      statVarRefList : "LKinLang_typeVarRefList";   // Table containing all variable references
      statLabelList : "LKinLang_typeLabelList";   // Table containing all label references
      statSubPrgList : "LKinLang_typeSubPrgList";   // Table containing all subprogram references
      statStack : "LKinLang_typeStack";   // Static storing for stack elements
      statHierarchicLevel : "LKInLang_typeHierarchicLevel";   // Static storing for hierarchic level info
   END_VAR
   VAR_TEMP
      tempExecute : Bool;   // Temporary value for input 'execute'
      tempStop : Bool;   // Temporary value for input 'stop'
      tempReturnVal : DWord;   // Temporary value for returns of functions
      tempError : Bool;   // Temporary value for error
      tempCounter : Int;   // Temporary counter variable
      tempLabelIndex : Int;   // Temporary counter in labelList
      tempEmptyLineCounter : Int;   // Temporary counter for empty lines / Tenporary counter for empty lines
      tempTokenCounter : Int;   // Temporary counter for token
      tempCycleCounter : Int;   // Temporary value for cycle counter
      tempParseCounter : Int;   // Temporary var to switch direct and follow value parsing
      tempFollowValueCounter : Int;   // Temporary counter for follow values
      tempConditionCounter : Int;   // Temporary counter for conditions
      tempWaitCheckCounter : Int;   // Temporary token counter to check for wait comamnds
      tempFlagOnly : Bool;   // Temporary bit to signalize flag only cmd
      tempWaitTime : Bool;   // Temporary bit to signalize a wait command
      tempAbortRepeat : Bool;   // Temporary bit to abort the repeat loop
      tempParameterIndex : Int;   // Temporary parameter index
      tempSeparatorIndex : Int;   // Temporary separator index
      tempCmdWord : Word;   // Temporary command word
      tempParameterValue : LReal;   // Temporary parameter value
      tempCmdName : String;   // Temporary command name
      tempVarType : Int;   // Temporary variable showing the type of a variable
      tempVarIndex : Int;   // Temporary variable showing the index of a variable
      tempLabelExists : Bool;   // Temporary bit to signalize if a label exists
      tempConditionResult : Bool;   // Temporary result of a condition for conditional jumps
      tempGlobal : Bool;   // Temporary bit to signalize a global variable
      tempPointerOk : Bool;   // Temporary bit to signalize line buffer pointer are ok
      tempLineNumber : UDInt;   // Temporary line number
      tempDelimPos : Array[1..3] of SInt;   // Temporary position of delimiters
      tempTestCommand : "LKinLang_typePathDataElement";   // Temporary PathData command to test iparsed is new
      tempParsedValues : "LKinCtrl_typePathDataElement_advanced";   // Temporary path data element with parsed values
      tempParameterCounter : Array[1.."LKINLANG_MAX_NUMBER_OF_PARAMETERS_PER_LINE"] of "LKinLang_typeParameterCounter";   // Counts the found parameter in one line (G1,F,...)
      tempWaitParameterDefinition : "LKinLang_typeParameterDefinition";   // Temporary definition for a wait command
      tempMathParserResult : "LKinLang_typeMathParserResult";   // Temporary result of the math parser
   END_VAR
   VAR CONSTANT
      MAX_LINES_PER_CYCLE : SInt := 1;   // Maximum lines to be parsed in one call
      MAX_EMPTY_LINES_PER_CYCLE : Int := 5;   // Maximum empty lines handled in one cycle
      MAX_LINES_LABEL_LIST : Int := 5;   // Maximum lines handled in one labelList cycle
      DEFAULT_FLAG_MODE : USInt := 1;   // Flag mode used, if no input default is set
      FB_STATE_NO_PROCESSING : DInt := 0;   // FB state: No processing
      FB_STATE_INIT : DInt := 10;   // FB state: Initialize
      FB_STATE_LOOKUP_PART_1 : DInt := 20;   // FB state: Get commands oart 1
      FB_STATE_LOOKUP_PART_2 : DInt := 21;   // FB state: Get commands part 2
      FB_STATE_PRECHECK_PRG : DInt := 22;   // FB state: Precheck program / FB state: Create label list
      FB_STATE_PARSING : DInt := 30;   // FB state: Parsing
      FB_STATE_STOPPING : DInt := 40;   // FB state: Stopping
      STATE_SEARCH_LINE : Int := 90;   // Internal FB state: Search line in buffer / Internal FB state: Wait until FileHandler has found requested line
      STATE_FILEHANDLER_REQUEST : Int := 91;   // Internal FB state: Wait until FileHandler has found requested line
      STATE_TOKENIZING : Int := 100;   // Internal FB state: Tokenizing
      STATE_INIT_PARSE_LINE : Int := 200;   // Internal FB state: Parsing
      STATE_IS_LINE_VAR_DEF : Int := 201;   // Internal FB state: Is line a variable definition
      STATE_LINE_IS_VAR_DEF : Int := 202;   // Internal FB state: Line is a variable definition
      STATE_IS_LINE_LABEL : Int := 203;   // Internal FB state: Is line a label
      STATE_IS_LINE_GOTO : Int := 204;   // Internal FB state: Is line is jump
      STATE_IS_LINE_STOPRE : Int := 205;   // Internal FB state: Is line a processing stop
      STATE_IS_LINE_IF : Int := 207;   // Internal FB state: Check if line contains IF
      STATE_IS_LINE_WHILE : Int := 208;   // Internal FB state: Check if line contains WHILE
      STATE_IS_LINE_FOR : Int := 209;   // Internal FB state: Check if line contains FOR
      STATE_IS_LINE_SUB : Int := 210;   // Internal FB state: Check if line contains SUB
      STATE_INIT_PARSE_LOOP : Int := 300;   // Internal FB state: Initialize parsing loop
      STATE_IS_TOKEN_SEPARATOR : Int := 310;   // Internal FB state: Check token for separator
      STATE_TOKEN_IS_SEPARATOR : Int := 311;   // Internal FB state: Token is separator
      STATE_IS_TOKEN_NUMBER : Int := 320;   // Internal FB state: Check token for number
      STATE_IS_TOKEN_PARAMETER : Int := 330;   // Internal FB state: Check token for parameter
      STATE_TOKEN_IS_PARAMETER : Int := 331;   // Internal FB state: Token is parameter
      STATE_IS_TOKEN_VARIABLE : Int := 340;   // Internal FB state: Check token for variable
      STATE_TOKEN_IS_VARIABLE : Int := 341;   // Internal FB state: Token is variable
      STATE_TOKEN_IS_UNKNOWN : Int := 350;   // Internal FB state: Token is unknown
      STATE_TOKEN_PROCESSED : Int := 390;   // Internal FB state: Token was processed
      STATE_LINE_PARSED : Int := 400;   // Internal FB state: Parsing single line done
      STATE_CHECK_FOR_NEW_PATH_DATA_CMD : Int := 500;   // Internal FB state: Check parsed command
      STATE_BUILD_PATH_DATA_CMD : Int := 600;   // Internal FB state: Build complete PathData command
      STATE_WRITE_CMD : Int := 700;   // Internal FB state: Write parsed command to path data
      STATE_RESET_AFTER_WRITE : Int := 701;   // Internal FB state: Reset statics and save "old" variables
      STATE_CHECK_END : Int := 800;   // Internal FB state: Check for end of program
      STATE_ERROR : Int := 900;   // Internal FB state: Error
      STATE_PREPROCESSING_STOP : Int := 1000;   // Internal FB state: Wait for MovePath to catch up with execution
      STATUS_EXECUTION_FINISHED : Word := 16#0000;   // Execution finished without errors
      STATUS_NO_CALL : Word := 16#7000;   // No job being currently processed
      STATUS_FIRST_CALL : Word := 16#7001;   // First call after incoming new job (rising edge 'execute')
      STATUS_SUBSEQUENT_CALL : Word := 16#7002;   // Subsequent call during active processing without further details
      STATUS_COMMAND_ABORTED : Word := 16#7FFF;   // Commanded functionality has been aborted by another command
      ERR_UNDEFINED_STATE : Word := 16#8600;   // Error due to an undefined state in state machine
      ERR_PARSING : Word := 16#8601;   // Error while parsing line
      ERR_TOKENIZING : Word := 16#8602;   // Error while tokenizing line
      ERR_LOOKUP : Word := 16#8603;   // Error while creating lookUp table
      ERR_HIERARCHIC_LEVEL_LIST : Word := 16#8604;   // Error while creating hierarchic level list
      ERR_LABEL_LIST : Word := 16#8605;   // Error while creating label list
      ERR_SUB_PROGRAM_LIST : Word := 16#8606;   // Error while creating sub program list
      ERR_LANGUAGE : Word := 16#8200;   // Error missing language definition
      ERR_WRONG_DEFAULTS : Int := -998;   // Error due to missing or wrong default connection
      ERR_LANG_NOT_DEFINED : Int := -999;   // Error selected language not defined
      MINVAL_LREAL : LReal := -1.7976931348623157E+308;   // Minimum value of LREAL
      MAXVAL_LREAL : LReal := 1.7976931348623157E+308;   // Minimum value of LREAL
      MINVAL_DINT : DInt := -2147483648 ;   // Minimum value of DINT
      MAXVAL_DINT : DInt := +2147483647;   // Minimum value of DINT
      MINVAL_INT : Int := -32768;   // Minimum value of INT
      MAXVAL_INT : Int := 32767;   // Maximum vlaue of INT
   END_VAR
BEGIN
   //==========================================================================================
   // SIEMENS AG
   // (c)Copyright 2020 All Rights Reserved
   //------------------------------------------------------------------------------------------
   // Library: LKinLang
   // Tested with: S7-1517T-3 PN/DP
   // Engineering: TIA Portal V15
   // Restrictions: ---
   // Requirements: S7-1500T FW 2.5
   // Functionality: LKinLang_Parser
   // The FB parses strings from line buffer to PathData commands using different language
   // packages.
   // 
   // Support: tech.team.motioncontrol@siemens.com
   // Note: Parameter comments are only available in language 'English (United States)'
   //------------------------------------------------------------------------------------------
   // Change log table:
   // Version    Date          Expert in charge    Changes applied
   // 01.00.00   28.05.2019    FR                  First created version
   // 01.00.01   16.07.2019    FR                  Fixed inserting relative cmd with length 0.0 in some unneccessary cases 
   // 01.00.02   29.07.2019    FR                  Reworked parsing; it is now done directly in this FB
   // 01.01.00   25.11.2019    FR                  Added LRealFlags
   //                                              Added FlagOnlyCmd
   //                                              Added default flag modes as input
   //                                              Fix ignoreAddPointer for LineBuffer
   // 01.01.01   12.02.2020    FR                  Fix circle (auxPoint) recognized as flagOnlyCmd
   // 01.01.02   17.02.2020    FR                  Fix for modal values not taken into account
   //                                              Changed transitionParameter[1] from Int to LReal
   // 01.01.03   17.02.2020    FR                  Changed approach to modal values
   // 01.02.00   15.04.2020    FR                  Added local variables, interface variables and jumps; Added remainingDistance to flagModeDefaults
   // 01.02.01   26.10.2020    FR                  Bugfix when generating label list
   // 01.03.00   01.12.2020    FR                  Added subprograms | Added IF,FOR,WHILE | Several bugfixes
   // 01.03.01   12.04.2021    FR                  Bugfix using followVal for circMode
   //===========================================================================================

   #tempExecute := #execute; // Work with temporary value / create process image
   #tempStop := #stop; // Work with temporary value / create process image

   REGION TRIGGERING
     IF #tempStop = TRUE AND (#statStopOld = FALSE) THEN
       // Stop FB execution
       #statFBState := #FB_STATE_STOPPING;
       // Set status here to avoid return in case of status = NO_CALL
       #statStatus := #STATUS_COMMAND_ABORTED;

     ELSIF (#tempExecute = TRUE) AND (#statExecuteOld = FALSE) AND (#tempStop = FALSE) // Check if FB is triggered
       AND (#statStatus = #STATUS_NO_CALL) // FB must be finished before new job can be started
     THEN // First call; initialize FB
       #statDone := FALSE;
       #statBusy := TRUE;
       #statCommandAborted := FALSE;
       #statError := FALSE;
       #statStatus := #STATUS_FIRST_CALL;

       // Init add pointer (path data)
       #statAddPointer := 0;
       #pathData.pointers.addPointer := 0;
       #pathData.pointers.bufferLocked := TRUE;
       #pathData.pointers.ignoreAddPointer := FALSE;
       #pathData.pointers.preprocessingStop := FALSE;

       // Init retrieve pointer to 0 (line buffer)
       #lineBuffer.pointers.retrievePointer := 0;

       // Reset Error String
       #statErrorString := '';

       // Init look up table
       FOR #tempCounter := 1 TO "LKINLANG_MAX_NUMBER_OF_PARAMETERS" DO
         #statParameterLookUpTable[#tempCounter].parameterNameString := '';
         #statParameterLookUpTable[#tempCounter].parameterNameNumber := 0;
         #statParameterLookUpTable[#tempCounter].parameterNumber := 0;
         #statParameterLookUpTable[#tempCounter].directValueWord := 16#0;
         FOR #tempFollowValueCounter := 1 TO "LKINLANG_NUMBER_OF_FOLLOW_VALUES" DO
           #statParameterLookUpTable[#tempCounter].followValueWords[#tempFollowValueCounter] := 16#0;
         END_FOR;
       END_FOR;

       // FR 2019/04/30
       // Reset path data 
       FOR #tempCounter := 1 TO "LKINCTRL_NO_OF_PATHDATA_ELEMENTS_ADVANCED" DO
         #pathData.commands[#tempCounter] := #statPathDataElementEmpty.pathDataElement;
       END_FOR;

       // Init empty path data element 
       #statModalCommand := #statPathDataElementEmpty;
       #statModalCommandOld := #statPathDataElementEmpty;
       #statModalProgram := #statPathDataElementEmpty;
       #statActualCommand := #statPathDataElementEmpty;
       #statActualCommandOld := #statPathDataElementEmpty;

       #statElementCounter := #statElementCounterEmpty;

       // Init conditions
       FOR #tempCounter := 1 TO "LKINLANG_NUMBER_OF_CONDITIONS" DO
         #statConditionsToCheck[#tempCounter] := #statConditionEmpty;
         #statSetParametersInCmd[#tempCounter] := #statConditionEmpty;
         #statSetParametersInPrg[#tempCounter] := #statConditionEmpty;
       END_FOR;

       // Init tokenized line
       #statTokenizedLine.lineNo := 0;
       #statTokenizedLine.numberOfToken := 0;
       FOR #tempCounter := 1 TO "LKINLANG_MAX_NUMBER_OF_TOKEN_PER_LINE" DO
         #statTokenizedLine.lineToken[#tempCounter] := '';
       END_FOR;

       // Init Positioning mode to absolute
       #statPositioningMode := 1;

       // Init token counter
       #tempTokenCounter := 1;

       // Init condition counter
       #tempConditionCounter := 1;

       // Init flag counter
       #statActualFlagNumber := 0;

       // Init variable definition
       #statVariableDeclaration.localVariables := '';
       #statVariableDeclaration.globalVariables := '';
       #statLocalVariableDefinition.tokenizedString.lineNo := 0;
       #statLocalVariableDefinition.tokenizedString.numberOfToken := 0;
       FOR #tempCounter := 1 TO "LKINLANG_MAX_NUMBER_OF_TOKEN_PER_LINE" DO
         #statLocalVariableDefinition.tokenizedString.lineToken[#tempCounter] := '';
       END_FOR;
       #statLocalVariableDefinition.nameTokenNumber := 0;
       #statLocalVariableDefinition.typeTokenNumber := 0;
       // Init global
       #statGlobalVariableDefinition := #statLocalVariableDefinition;


       // Init vars & counter
       FOR #tempVarIndex := 1 TO "LKINLANG_NUMBER_OF_LOCAL_BOOL" DO
         #statVariables.boolean[#tempVarIndex] := FALSE;
       END_FOR;
       FOR #tempVarIndex := 1 TO "LKINLANG_NUMBER_OF_LOCAL_DINT" DO
         #statVariables.dints[#tempVarIndex] := 0;
       END_FOR;
       FOR #tempVarIndex := 1 TO "LKINLANG_NUMBER_OF_LOCAL_LREAL" DO
         #statVariables.lreals[#tempVarIndex] := 0.0;
       END_FOR;
       #statVariables.boolCounter := 0;
       #statVariables.dintCounter := 0;
       #statVariables.lrealCounter := 0;

       // Remove local vars from var ref table
       FOR #tempVarIndex := 1 TO "LKINLANG_NUMBER_OF_VAR_REFS" DO
         IF #statVarRefList.references[#tempVarIndex].type < "LKINLANG_VAR_TYPE_INTERFACE_BOOL" THEN
           #statVarRefList.references[#tempVarIndex].index := 0;
           #statVarRefList.references[#tempVarIndex].name := '';
           #statVarRefList.references[#tempVarIndex].type := 0;
           #statVarRefList.references[#tempVarIndex].scope := 0;
         END_IF;
       END_FOR;

       // Reset number of references
       #statVarRefList.numberOfReferences := 0;

       // Reset LabelList
       FOR #tempCounter := 1 TO "LKINLANG_NUMBER_OF_LABELS" DO
         #statLabelList.labels[#tempCounter].labelName := '';
         #statLabelList.labels[#tempCounter].lineNumber := 0;
         #statLabelList.labels[#tempCounter].hierarchicLevel := 0;
       END_FOR;
       #statLabelList.numberOfLabels := 0;

       // Reset hierarchicLevel
       FOR #tempCounter := 1 TO "LKINLANG_NUMBER_OF_HIERARCHICLEVEL" DO
         #statHierarchicLevel.levels[#tempCounter].level := 0;
         #statHierarchicLevel.levels[#tempCounter].lineNumber := 0;
         #statHierarchicLevel.levels[#tempCounter].type := 0;
       END_FOR;
       #statHierarchicLevel.numberOfLevels := 0;
       #statHierarchicLevel.currentLevel := 0;

       // Reset Stack
       FOR #tempCounter := 1 TO "LKINLANG_NUMBER_OF_STACK_ELEMENTS" DO
         #statStack.stackElements[#tempCounter].lineNumberStart := 0;
         #statStack.stackElements[#tempCounter].lineNumberEnd := 0;
         #statStack.stackElements[#tempCounter].type := 0;
         #statStack.stackElements[#tempCounter].increment := 0;
         #statStack.stackElements[#tempCounter].quantity := 0;
         #statStack.stackElements[#tempCounter].variableRef.index := 0;
         #statStack.stackElements[#tempCounter].variableRef.type := 0;
         #statStack.stackElements[#tempCounter].variableRef.name := '';
       END_FOR;
       #statStack.numberOfElements := 0;

       // Reset subprogram list
       FOR #tempCounter := 1 TO "LKINLANG_NUMBER_OF_SUBPROGRAMS" DO
         #statSubPrgList.subPrgs[#tempCounter].prgName := '';
         #statSubPrgList.subPrgs[#tempCounter].lineNumberStart := 0;
         #statSubPrgList.subPrgs[#tempCounter].lineNumberEnd := 0;
       END_FOR;
       #statSubPrgList.numberOfSubPrgs := 0;

       // Reset parameter definition
       #statParameterDefinition := #statParameterDefinitionEmpty;

       // Select Language
       #statSelectedLanguage := #language;

       // Syntax check
       #statSyntaxCheck := #syntaxCheck;

       // Reset stringExpression
       #statStringExpression := '';

       // Reset requested line
       #statSearchedLine := 0;

       // Set file state initially
       IF #lineBuffer.info.fileState = "LKINLANG_FILE_STATE_LOADING" THEN
         #lineBuffer.info.fileState := "LKINLANG_FILE_STATE_RUNNING_LOADING";
       ELSE
         #lineBuffer.info.fileState := "LKINLANG_FILE_STATE_RUNNING";
       END_IF;

       // State machine - start processing
       #statFBState := #FB_STATE_INIT;

     ELSIF (#statStatus = #STATUS_FIRST_CALL) THEN
       #statStatus := #STATUS_SUBSEQUENT_CALL;
     END_IF;

     // Edge detection 'execute' input
     #statExecuteOld := #tempExecute;
     // Edge detection 'stop' input
     #statStopOld := #tempStop;
   END_REGION TRIGGERING

   IF (#statStatus = #STATUS_NO_CALL) THEN // Nothing to do -> End here to reduce "system load"
     RETURN;
   END_IF;

   REGION STATE_MACHINE
     CASE #statFBState OF // State machine of FB
       #FB_STATE_NO_PROCESSING: // No processing active (Note: this state must always be present and left empty)
         ;

         // ------------------------------------------------------------------------------------------
         // Get separators, mergers and valid counts from language and save in static arrays
         // ------------------------------------------------------------------------------------------  
       #FB_STATE_INIT:
         REGION FB_STATE_INIT
           // Get separators and mergers from language package
           #tempParameterIndex := -1;
           "LKinLang_SelectLangPackage"(language := #statSelectedLanguage,
                                        variableDeclarations => #statVariableDeclaration,
                                        keyToken => #statKeyToken,
                                        parameterDefinition := #statParameterDefinition,
                                        separators => #statSeparators,
                                        mergers => #statMergers,
                                        validCounts => #statValidCounts,
                                        parameterNumber := #tempParameterIndex,
                                        parameterDefaults := #parameterDefaults);

           IF #tempParameterIndex = #ERR_LANG_NOT_DEFINED THEN
             // Error language not defined
             #statStatus := #ERR_LANGUAGE;
             #statStateIntern := #STATE_ERROR;
             #statErrorString := CONCAT(IN1 := #statErrorString, IN2 := 'Error: Selected language ');
             #statErrorString := CONCAT(IN1 := #statErrorString, IN2 := INT_TO_STRING(#statSelectedLanguage));
             #statErrorString := CONCAT(IN1 := #statErrorString, IN2 := ' not defined');
           END_IF;

           IF #tempParameterIndex = #ERR_WRONG_DEFAULTS THEN
             // Error language not defined
             #statStatus := #ERR_LANGUAGE;
             #statStateIntern := #STATE_ERROR;
             #statErrorString := CONCAT(IN1 := #statErrorString, IN2 := 'Error: Type of parameter defaults not matching language');
           END_IF;

           #statLastIndexOfMerger := 1;

           // Search last entry in mergers to save time in tokenizing
           FOR #tempCounter := 1 TO "LKINLANG_NUMBER_OF_MERGERS" DO
             IF #statMergers[#tempCounter] <> 16#00 THEN
               #statLastIndexOfMerger := #tempCounter;
             END_IF;
           END_FOR;

           // Tokenize variable definition string from language package
           #tempReturnVal := "LKinLang_TokenizeSlot"(lastIndexOfMerger := #statLastIndexOfMerger,
                                                     lineNumber := 0,
                                                     line := #statVariableDeclaration.localVariables,
                                                     separators := #statSeparators,
                                                     mergers := #statMergers,
                                                     preprocessorConfig := #preProcessConfig,
                                                     tokenizedLine => #statLocalVariableDefinition.tokenizedString,
                                                     errorString := #statErrorString);

           // Search tokenized variable definiton for name and type token
           FOR #tempCounter := 1 TO #statLocalVariableDefinition.tokenizedString.numberOfToken DO
             IF #statLocalVariableDefinition.tokenizedString.lineToken[#tempCounter] = '_name_' THEN
               #statLocalVariableDefinition.nameTokenNumber := DINT_TO_USINT(#tempCounter);
             ELSIF #statLocalVariableDefinition.tokenizedString.lineToken[#tempCounter] = '_type_' THEN
               #statLocalVariableDefinition.typeTokenNumber := DINT_TO_USINT(#tempCounter);
             END_IF;
           END_FOR;

           // Double check 
           IF #statLocalVariableDefinition.nameTokenNumber = 0
             OR #statLocalVariableDefinition.typeTokenNumber = 0 THEN
             // Error no valid variable definition found
             #statStatus := #ERR_LANGUAGE;
             #statStateIntern := #STATE_ERROR;
             #statErrorString := CONCAT(IN1 := #statErrorString, IN2 := 'Error: No valid variable definition found');
           END_IF;

           // Tokenize variable definition string from language package
           #tempReturnVal := "LKinLang_TokenizeSlot"(lastIndexOfMerger := #statLastIndexOfMerger,
                                                     lineNumber := 0,
                                                     line := #statVariableDeclaration.globalVariables,
                                                     separators := #statSeparators,
                                                     mergers := #statMergers,
                                                     preprocessorConfig := #preProcessConfig,
                                                     tokenizedLine => #statGlobalVariableDefinition.tokenizedString,
                                                     errorString := #statErrorString);

           // Search tokenized variable definiton for name and type token
           FOR #tempCounter := 1 TO #statGlobalVariableDefinition.tokenizedString.numberOfToken DO
             IF #statGlobalVariableDefinition.tokenizedString.lineToken[#tempCounter] = '_name_' THEN
               #statGlobalVariableDefinition.nameTokenNumber := DINT_TO_USINT(#tempCounter);
             ELSIF #statGlobalVariableDefinition.tokenizedString.lineToken[#tempCounter] = '_type_' THEN
               #statGlobalVariableDefinition.typeTokenNumber := DINT_TO_USINT(#tempCounter);
             END_IF;
           END_FOR;

           // Double check 
           IF #statGlobalVariableDefinition.nameTokenNumber = 0
             OR #statGlobalVariableDefinition.typeTokenNumber = 0 THEN
             // Error no valid variable definition found
             #statStatus := #ERR_LANGUAGE;
             #statStateIntern := #STATE_ERROR;
             #statErrorString := CONCAT(IN1 := #statErrorString, IN2 := 'Error: No valid variable definition found');
           END_IF;

           // Check syntax check mode
           IF #statSyntaxCheck <> "LKINLANG_SYNTAX_CHECK_AND_EXECUTE"
             AND #statSyntaxCheck <> "LKINLANG_SYNTAX_CHECK_OFF"
             AND #statSyntaxCheck <> "LKINLANG_SYNTAX_CHECK_ONLY" THEN
             // Error no valid syntax check mode
             #statStatus := #ERR_LANGUAGE;
             #statStateIntern := #STATE_ERROR;
             #statErrorString := CONCAT(IN1 := #statErrorString, IN2 := 'Error: No valid syntax check setting');
           END_IF;

           // Next state
           #statFBState := #FB_STATE_LOOKUP_PART_1;
         END_REGION FB_STATE_INIT

         // ------------------------------------------------------------------------------------------
         // Get first part of language definition where ParameterNameNumber <> -1 
         // Save the parameter numbers in lookup-table
         // The lookup-table is later used while parsing to have faster access to the parameter definition
         // ------------------------------------------------------------------------------------------ 
       #FB_STATE_LOOKUP_PART_1:
         REGION FB_STATE_LOOKUP_PART_1
           // Init command counter
           #statLookUpTableCounter := 1;

           // Get commands with parameterNameNumber <> -1
           "LKinLang_CreateParameterLookUpTable"(language := #statSelectedLanguage,
                                                 mode := 0, //  ParameterNameNumber <> -1
                                                 error => #tempError,
                                                 lastIndexLookUp => #statLastIndexLookUp,
                                                 parameterLookUpTable := #statParameterLookUpTable,
                                                 parameterDefaults := #parameterDefaults,
                                                 parameterCounter := #statLookUpTableCounter,
                                                 errorString := #statErrorString);
           IF #tempError THEN
             // Error while creating look up table --> Exit
             #statStatus := #ERR_LOOKUP;
             #statStateIntern := #STATE_ERROR;
           ELSE
             // Next state
             #statFBState := #FB_STATE_LOOKUP_PART_2;
           END_IF;
         END_REGION FB_STATE_LOOKUP_PART_1

         // ------------------------------------------------------------------------------------------
         // Get second part of language definition where ParameterNameNumber = -1 
         // Save the parameter numbers in lookup-table
         // Initialize internal states (IF cases)
         // ------------------------------------------------------------------------------------------ 
       #FB_STATE_LOOKUP_PART_2:
         REGION FB_STATE_LOOKUP_PART_2
           // Get commands with parameterNameNumber = -1
           "LKinLang_CreateParameterLookUpTable"(language := #statSelectedLanguage,
                                                 mode := 1, // ParameterNameNumber = -1
                                                 error => #tempError,
                                                 lastIndexLookUp => #statLastIndexLookUp,
                                                 parameterLookUpTable := #statParameterLookUpTable,
                                                 parameterDefaults := #parameterDefaults,
                                                 parameterCounter := #statLookUpTableCounter,
                                                 errorString := #statErrorString);
           IF #tempError THEN
             // Error while creating look up table --> Exit
             #statStatus := #ERR_LOOKUP;
             #statStateIntern := #STATE_ERROR;
           ELSE
             // Next state
             //#statFBState := #FB_STATE_PARSING;
             #statFBState := #FB_STATE_PRECHECK_PRG;

             // Set internal state to tokenizing
             #statStateIntern := #STATE_TOKENIZING;
           END_IF;
         END_REGION FB_STATE_LOOKUP_PART_2

         // ------------------------------------------------------------------------------------------
         // Here the whole program is checked
         // Following things should be done here:
         // - Get HierarchicLevel
         // - Create Label List
         // - Get ProgramName (PRG)?
         // - Get SubProgram List
         // - Check for M17/M30?
         //  
         // After all this is done without error, the actual parsing can be started 
         // The filehandler must be restarted and the lineBuffer must be reset
         // then switch over to FB state "PARSING"
         // The tokenization has to be done here and in state PARSING --> Maybe find a better solution?
         // ------------------------------------------------------------------------------------------
       #FB_STATE_PRECHECK_PRG:
         REGION FB_STATE_PRECHECK_PRG
           // Reset empty line counter
           #tempEmptyLineCounter := 0;

           // Repeat tokenizing until aborted
           // Aborted by:
           // - No new lines in line buffer
           // - End of file reached
           REPEAT

             // Check lineBuffer pointer if next line can be retrieved
             IF ((#lineBuffer.pointers.addPointer > #lineBuffer.pointers.retrievePointer
               AND NOT #lineBuffer.pointers.bufferLocked // Buffer is not locked by fileHandler
               AND NOT #lineBuffer.pointers.addPointerRestarted) // Overflow of ring buffer
               OR
               (#lineBuffer.pointers.addPointer < #lineBuffer.pointers.retrievePointer
               AND #lineBuffer.pointers.addPointerRestarted
               AND NOT #lineBuffer.pointers.bufferLocked))
               OR #lineBuffer.pointers.ignoreAddPointer // FR 25.11.2019
             THEN

               // Increment retrieve pointer
               IF #lineBuffer.pointers.retrievePointer < "LKINLANG_LAST_INDEX_LINE_BUFFER" THEN
                 #lineBuffer.pointers.retrievePointer += 1;

                 // Reset retrieve pointer to 1 and reset overflow variable
               ELSIF #lineBuffer.pointers.retrievePointer >= "LKINLANG_LAST_INDEX_LINE_BUFFER" THEN
                 #lineBuffer.pointers.retrievePointer := 1;
                 #lineBuffer.pointers.addPointerRestarted := FALSE;
               END_IF;

               // ------------------------------------------------------------------------------------------
               // Get hierarchic level
               // ------------------------------------------------------------------------------------------
               // Get hierarchic level --> Check for IF;WHILE;FOR and increse or decrease level
               // Hierarchic level is needed to check if jumps are allowed
               REGION GET_HIERARCHIC_LEVEL
                 // Check if line contains IF token
                 IF FIND(IN1 := #lineBuffer.lines[#lineBuffer.pointers.retrievePointer].content, IN2 := #statKeyToken.tokenIf) <> 0 THEN
                   // Tokenize line where retrieve pointer is pointing at
                   #tempReturnVal := "LKinLang_TokenizeSlot"(lastIndexOfMerger := #statLastIndexOfMerger,
                                                             lineNumber := #lineBuffer.lines[#lineBuffer.pointers.retrievePointer].number,
                                                             line := #lineBuffer.lines[#lineBuffer.pointers.retrievePointer].content,
                                                             separators := #statSeparators,
                                                             mergers := #statMergers,
                                                             preprocessorConfig := #preProcessConfig,
                                                             tokenizedLine => #statTokenizedLine,
                                                             errorString := #statErrorString);

                   // Check if line has content
                   IF #statTokenizedLine.numberOfToken > 0 THEN
                     // Check if line starts with IF token
                     IF #statTokenizedLine.lineToken[#statTokenizedLine.numberOfToken] = #statKeyToken.tokenIf THEN
                       // Increase array index
                       #statHierarchicLevel.numberOfLevels += 1;
                       // Check if index is ok
                       IF #statHierarchicLevel.numberOfLevels <= "LKINLANG_NUMBER_OF_HIERARCHICLEVEL" THEN
                         // Increase hierarchic level
                         #statHierarchicLevel.currentLevel += 1;
                         // Store entry
                         #statHierarchicLevel.levels[#statHierarchicLevel.numberOfLevels].level := #statHierarchicLevel.currentLevel;
                         #statHierarchicLevel.levels[#statHierarchicLevel.numberOfLevels].lineNumber := #statTokenizedLine.lineNo;
                         #statHierarchicLevel.levels[#statHierarchicLevel.numberOfLevels].type := "LKINLANG_ENTRY_TYPE_IF"; // Type for IF
                       ELSE
                         // Error hierarchic level array overflow
                         #statStatus := #ERR_HIERARCHIC_LEVEL_LIST;
                         #statStateIntern := #STATE_ERROR;
                         #statErrorString := CONCAT(IN1 := #statErrorString, IN2 := 'Error: Maximum array index of hierarchic level reached');
                         #statErrorString := CONCAT(IN1 := #statErrorString, IN2 := ' in line: ');
                         #statErrorString := CONCAT(IN1 := #statErrorString, IN2 := UDINT_TO_STRING(#statTokenizedLine.lineNo));
                       END_IF;
                     END_IF;
                   END_IF;
                 END_IF;

                 // Check if line contains ELSE token
                 IF FIND(IN1 := #lineBuffer.lines[#lineBuffer.pointers.retrievePointer].content, IN2 := #statKeyToken.tokenElse) <> 0 THEN
                   // Tokenize line where retrieve pointer is pointing at
                   #tempReturnVal := "LKinLang_TokenizeSlot"(lastIndexOfMerger := #statLastIndexOfMerger,
                                                             lineNumber := #lineBuffer.lines[#lineBuffer.pointers.retrievePointer].number,
                                                             line := #lineBuffer.lines[#lineBuffer.pointers.retrievePointer].content,
                                                             separators := #statSeparators,
                                                             mergers := #statMergers,
                                                             preprocessorConfig := #preProcessConfig,
                                                             tokenizedLine => #statTokenizedLine,
                                                             errorString := #statErrorString);

                   // Check if line has content
                   IF #statTokenizedLine.numberOfToken > 0 THEN
                     // Check if line starts with ELSE token
                     IF #statTokenizedLine.lineToken[#statTokenizedLine.numberOfToken] = #statKeyToken.tokenElse THEN
                       // Check if number of token is exactly 1 --> Nothing more allowed
                       IF #statTokenizedLine.numberOfToken = 1 THEN
                         // Increase array index
                         #statHierarchicLevel.numberOfLevels += 1;
                         // Check if index is ok
                         IF #statHierarchicLevel.numberOfLevels <= "LKINLANG_NUMBER_OF_HIERARCHICLEVEL" THEN
                           // Level does not change
                           // Store entry
                           #statHierarchicLevel.levels[#statHierarchicLevel.numberOfLevels].level := #statHierarchicLevel.currentLevel;
                           #statHierarchicLevel.levels[#statHierarchicLevel.numberOfLevels].lineNumber := #statTokenizedLine.lineNo;
                           #statHierarchicLevel.levels[#statHierarchicLevel.numberOfLevels].type := "LKINLANG_ENTRY_TYPE_ELSE"; // Type for ELSE
                         ELSE
                           // Error hierarchic level array overflow
                           #statStatus := #ERR_HIERARCHIC_LEVEL_LIST;
                           #statStateIntern := #STATE_ERROR;
                           #statErrorString := CONCAT(IN1 := #statErrorString, IN2 := 'Error: Maximum array index of hierarchic level reached');
                           #statErrorString := CONCAT(IN1 := #statErrorString, IN2 := ' in line: ');
                           #statErrorString := CONCAT(IN1 := #statErrorString, IN2 := UDINT_TO_STRING(#statTokenizedLine.lineNo));
                         END_IF;
                       ELSE
                         // Error wrong usage of ELSE
                         #statStatus := #ERR_HIERARCHIC_LEVEL_LIST;
                         #statStateIntern := #STATE_ERROR;
                         #statErrorString := CONCAT(IN1 := #statErrorString, IN2 := 'Error: Wrong syntax of ');
                         #statErrorString := CONCAT(IN1 := #statErrorString, IN2 := #statKeyToken.tokenElse);
                         #statErrorString := CONCAT(IN1 := #statErrorString, IN2 := ' in line: ');
                         #statErrorString := CONCAT(IN1 := #statErrorString, IN2 := UDINT_TO_STRING(#statTokenizedLine.lineNo));
                       END_IF;
                     END_IF;
                   END_IF;
                 END_IF;

                 // Check if line contains ENDIF token
                 IF FIND(IN1 := #lineBuffer.lines[#lineBuffer.pointers.retrievePointer].content, IN2 := #statKeyToken.tokenEndIf) <> 0 THEN
                   // Tokenize line where retrieve pointer is pointing at
                   #tempReturnVal := "LKinLang_TokenizeSlot"(lastIndexOfMerger := #statLastIndexOfMerger,
                                                             lineNumber := #lineBuffer.lines[#lineBuffer.pointers.retrievePointer].number,
                                                             line := #lineBuffer.lines[#lineBuffer.pointers.retrievePointer].content,
                                                             separators := #statSeparators,
                                                             mergers := #statMergers,
                                                             preprocessorConfig := #preProcessConfig,
                                                             tokenizedLine => #statTokenizedLine,
                                                             errorString := #statErrorString);

                   // Check if line has content
                   IF #statTokenizedLine.numberOfToken > 0 THEN
                     // Check if line starts with ENDIF token
                     IF #statTokenizedLine.lineToken[#statTokenizedLine.numberOfToken] = #statKeyToken.tokenEndIf THEN
                       // Check if number of token is exactly 1 --> Nothing more allowed
                       IF #statTokenizedLine.numberOfToken = 1 THEN
                         // Increase array index
                         #statHierarchicLevel.numberOfLevels += 1;
                         // Check if index is ok
                         IF #statHierarchicLevel.numberOfLevels <= "LKINLANG_NUMBER_OF_HIERARCHICLEVEL" THEN
                           // Store entry
                           #statHierarchicLevel.levels[#statHierarchicLevel.numberOfLevels].level := #statHierarchicLevel.currentLevel;
                           #statHierarchicLevel.levels[#statHierarchicLevel.numberOfLevels].lineNumber := #statTokenizedLine.lineNo;
                           #statHierarchicLevel.levels[#statHierarchicLevel.numberOfLevels].type := "LKINLANG_ENTRY_TYPE_ENDIF"; // Type for ENDIF

                           // Decrease hierarchic level
                           #statHierarchicLevel.currentLevel -= 1;
                         ELSE
                           // Error hierarchic level array overflow
                           #statStatus := #ERR_HIERARCHIC_LEVEL_LIST;
                           #statStateIntern := #STATE_ERROR;
                           #statErrorString := CONCAT(IN1 := #statErrorString, IN2 := 'Error: Maximum array index of hierarchic level reached');
                           #statErrorString := CONCAT(IN1 := #statErrorString, IN2 := ' in line: ');
                           #statErrorString := CONCAT(IN1 := #statErrorString, IN2 := UDINT_TO_STRING(#statTokenizedLine.lineNo));
                         END_IF;
                       ELSE
                         // Error wrong usage of ENDIF
                         #statStatus := #ERR_HIERARCHIC_LEVEL_LIST;
                         #statStateIntern := #STATE_ERROR;
                         #statErrorString := CONCAT(IN1 := #statErrorString, IN2 := 'Error: Wrong syntax of ');
                         #statErrorString := CONCAT(IN1 := #statErrorString, IN2 := #statKeyToken.tokenEndIf);
                         #statErrorString := CONCAT(IN1 := #statErrorString, IN2 := ' in line: ');
                         #statErrorString := CONCAT(IN1 := #statErrorString, IN2 := UDINT_TO_STRING(#statTokenizedLine.lineNo));
                       END_IF;
                     END_IF;
                   END_IF;
                 END_IF;

                 // Check if line contains WHILE token
                 IF FIND(IN1 := #lineBuffer.lines[#lineBuffer.pointers.retrievePointer].content, IN2 := #statKeyToken.tokenWhile) <> 0 THEN
                   // Tokenize line where retrieve pointer is pointing at
                   #tempReturnVal := "LKinLang_TokenizeSlot"(lastIndexOfMerger := #statLastIndexOfMerger,
                                                             lineNumber := #lineBuffer.lines[#lineBuffer.pointers.retrievePointer].number,
                                                             line := #lineBuffer.lines[#lineBuffer.pointers.retrievePointer].content,
                                                             separators := #statSeparators,
                                                             mergers := #statMergers,
                                                             preprocessorConfig := #preProcessConfig,
                                                             tokenizedLine => #statTokenizedLine,
                                                             errorString := #statErrorString);

                   // Check if line has content
                   IF #statTokenizedLine.numberOfToken > 0 THEN
                     // Check if line starts with WHILE token
                     IF #statTokenizedLine.lineToken[#statTokenizedLine.numberOfToken] = #statKeyToken.tokenWhile THEN
                       // Increase array index
                       #statHierarchicLevel.numberOfLevels += 1;
                       // Check if index is ok
                       IF #statHierarchicLevel.numberOfLevels <= "LKINLANG_NUMBER_OF_HIERARCHICLEVEL" THEN
                         // Increase hierarchic level
                         #statHierarchicLevel.currentLevel += 1;
                         // Store entry
                         #statHierarchicLevel.levels[#statHierarchicLevel.numberOfLevels].level := #statHierarchicLevel.currentLevel;
                         #statHierarchicLevel.levels[#statHierarchicLevel.numberOfLevels].lineNumber := #statTokenizedLine.lineNo;
                         #statHierarchicLevel.levels[#statHierarchicLevel.numberOfLevels].type := "LKINLANG_ENTRY_TYPE_WHILE"; // Type for WHILE
                       ELSE
                         // Error hierarchic level array overflow
                         #statStatus := #ERR_HIERARCHIC_LEVEL_LIST;
                         #statStateIntern := #STATE_ERROR;
                         #statErrorString := CONCAT(IN1 := #statErrorString, IN2 := 'Error: Maximum array index of hierarchic level reached');
                         #statErrorString := CONCAT(IN1 := #statErrorString, IN2 := ' in line: ');
                         #statErrorString := CONCAT(IN1 := #statErrorString, IN2 := UDINT_TO_STRING(#statTokenizedLine.lineNo));
                       END_IF;
                     END_IF;
                   END_IF;
                 END_IF;

                 // Check if line contains ENDWHILE token
                 IF FIND(IN1 := #lineBuffer.lines[#lineBuffer.pointers.retrievePointer].content, IN2 := #statKeyToken.tokenEndWhile) <> 0 THEN
                   // Tokenize line where retrieve pointer is pointing at
                   #tempReturnVal := "LKinLang_TokenizeSlot"(lastIndexOfMerger := #statLastIndexOfMerger,
                                                             lineNumber := #lineBuffer.lines[#lineBuffer.pointers.retrievePointer].number,
                                                             line := #lineBuffer.lines[#lineBuffer.pointers.retrievePointer].content,
                                                             separators := #statSeparators,
                                                             mergers := #statMergers,
                                                             preprocessorConfig := #preProcessConfig,
                                                             tokenizedLine => #statTokenizedLine,
                                                             errorString := #statErrorString);

                   // Check if line has content
                   IF #statTokenizedLine.numberOfToken > 0 THEN
                     // Check if line starts with ENDWHILE token
                     IF #statTokenizedLine.lineToken[#statTokenizedLine.numberOfToken] = #statKeyToken.tokenEndWhile THEN
                       // Check if number of token is exactly 1 --> Nothing more allowed
                       IF #statTokenizedLine.numberOfToken = 1 THEN
                         // Increase array index
                         #statHierarchicLevel.numberOfLevels += 1;
                         // Check if index is ok
                         IF #statHierarchicLevel.numberOfLevels <= "LKINLANG_NUMBER_OF_HIERARCHICLEVEL" THEN
                           // Store entry
                           #statHierarchicLevel.levels[#statHierarchicLevel.numberOfLevels].level := #statHierarchicLevel.currentLevel;
                           #statHierarchicLevel.levels[#statHierarchicLevel.numberOfLevels].lineNumber := #statTokenizedLine.lineNo;
                           #statHierarchicLevel.levels[#statHierarchicLevel.numberOfLevels].type := "LKINLANG_ENTRY_TYPE_ENDWHILE"; // Type for ENDWHILE

                           // Decrease hierarchic level
                           #statHierarchicLevel.currentLevel -= 1;
                         ELSE
                           // Error hierarchic level array overflow
                           #statStatus := #ERR_HIERARCHIC_LEVEL_LIST;
                           #statStateIntern := #STATE_ERROR;
                           #statErrorString := CONCAT(IN1 := #statErrorString, IN2 := 'Error: Maximum array index of hierarchic level reached');
                           #statErrorString := CONCAT(IN1 := #statErrorString, IN2 := ' in line: ');
                           #statErrorString := CONCAT(IN1 := #statErrorString, IN2 := UDINT_TO_STRING(#statTokenizedLine.lineNo));
                         END_IF;
                       ELSE
                         // Error wrong usage of ENDWHILE
                         #statStatus := #ERR_HIERARCHIC_LEVEL_LIST;
                         #statStateIntern := #STATE_ERROR;
                         #statErrorString := CONCAT(IN1 := #statErrorString, IN2 := 'Error: Wrong syntax of ');
                         #statErrorString := CONCAT(IN1 := #statErrorString, IN2 := #statKeyToken.tokenEndWhile);
                         #statErrorString := CONCAT(IN1 := #statErrorString, IN2 := ' in line: ');
                         #statErrorString := CONCAT(IN1 := #statErrorString, IN2 := UDINT_TO_STRING(#statTokenizedLine.lineNo));
                       END_IF;
                     END_IF;
                   END_IF;
                 END_IF;

